(* Logix 5000 project; controller FV vendor 1 type 14 code 217 rev 31.11; software revision 31.00; part 19 of 63 *)
(* tags used below, declared in another part *)
   CheckTimeMask : INT;
   Delphi_Does_Eng_Func : BOOL;
   FR_FRV1_AV01 : PlantItem;   // FRV1_AV01
   FR_FV26_AV01 : PlantItem;   // FV26_AV01
   FR_FV26_AV04 : PlantItem;   // FV26_AV04
   FR_FV28_VA01 : PlantItem;   // FV28_VA01
   FR_FV29_VA01 : PlantItem;   // FV29_VA01
   FR_FV30_VA01 : PlantItem;   // FV30_VA01
   FR_FV31_VA01 : PlantItem;   // FV31_VA01
   FR_FVR1_P01 : PlantItem;   // FVR1_P01
   FR_FVS_P01 : PlantItem;   // FVS_P01
   FR_GBM_P01 : PlantItem;   // GBM_P01
   FR_N255 : INT[265];   // CHECKWORDS
   FR_YM_P01 : PlantItem;   // YM_P01
   FR_YM_P02 : PlantItem;   // YM_P02
   FR_YM_P03 : PlantItem;   // YM_P03
   TempChecktime : DINT;
(* FR_Common, continued *)

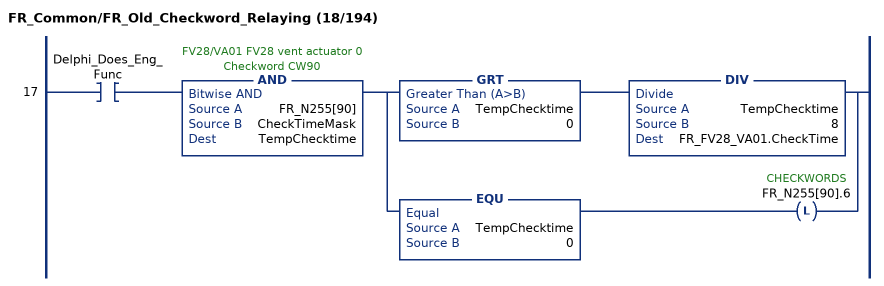
   [picture p322: FR_Common/FR_Old_Checkword_Relaying rungs 17-17]
   17: XIC(Delphi_Does_Eng_Func)AND(FR_N255[90],CheckTimeMask,TempChecktime)[GRT(TempChecktime,0) DIV(TempChecktime,8,FR_FV28_VA01.CheckTime) ,EQU(TempChecktime,0) OTL(FR_N255[90].6) ];
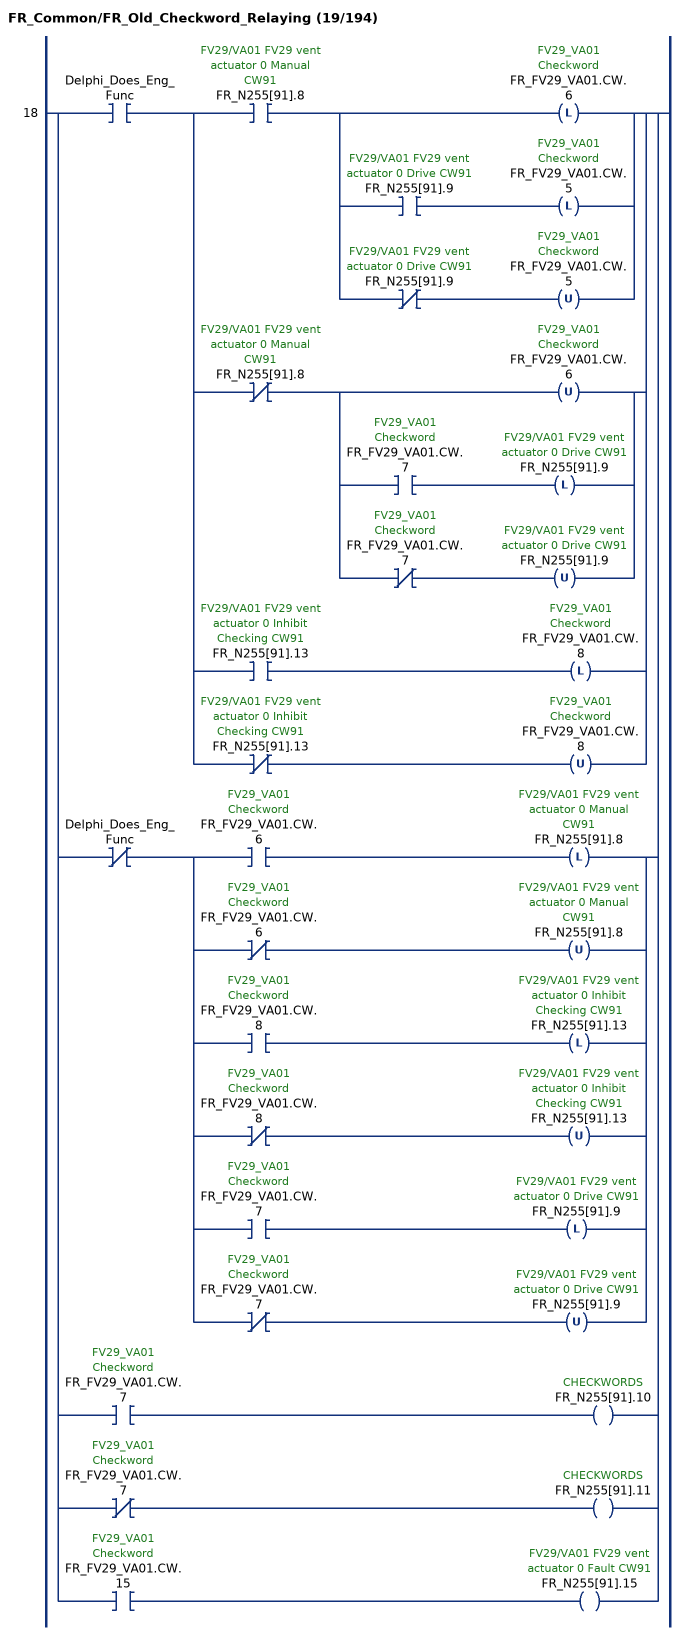
   18: [XIC(Delphi_Does_Eng_Func) [[XIC(FR_N255[91].8) [OTL(FR_FV29_VA01.CW.6) ,XIC(FR_N255[91].9) OTL(FR_FV29_VA01.CW.5) ,XIO(FR_N255[91].9) OTU(FR_FV29_VA01.CW.5) ] ,XIO(FR_N255[91].8) [OTU(FR_FV29_VA01.CW.6) ,[XIC(FR_FV29_VA01.CW.7) OTL(FR_N255[91].9) ,XIO(FR_FV29_VA01.CW.7) OTU(FR_N255[91].9) ] ] ] ,[XIC(FR_N255[91].13) OTL(FR_FV29_VA01.CW.8) ,XIO(FR_N255[91].13) OTU(FR_FV29_VA01.CW.8) ] ] ,XIO(Delphi_Does_Eng_Func) [[XIC(FR_FV29_VA01.CW.6) OTL(FR_N255[91].8) ,XIO(FR_FV29_VA01.CW.6) OTU(FR_N255[91].8) ] ,[XIC(FR_FV29_VA01.CW.8) OTL(FR_N255[91].13) ,XIO(FR_FV29_VA01.CW.8) OTU(FR_N255[91].13) ] ,[XIC(FR_FV29_VA01.CW.7) OTL(FR_N255[91].9) ,XIO(FR_FV29_VA01.CW.7) OTU(FR_N255[91].9) ] ] ,XIC(FR_FV29_VA01.CW.7) OTE(FR_N255[91].10) ,XIO(FR_FV29_VA01.CW.7) OTE(FR_N255[91].11) ,XIC(FR_FV29_VA01.CW.15) OTE(FR_N255[91].15) ];
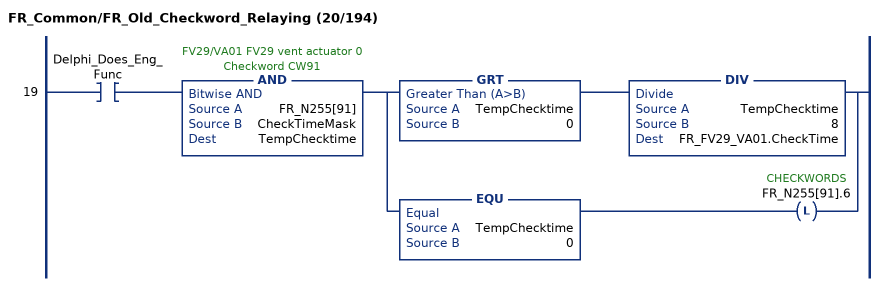
   19: XIC(Delphi_Does_Eng_Func)AND(FR_N255[91],CheckTimeMask,TempChecktime)[GRT(TempChecktime,0) DIV(TempChecktime,8,FR_FV29_VA01.CheckTime) ,EQU(TempChecktime,0) OTL(FR_N255[91].6) ];
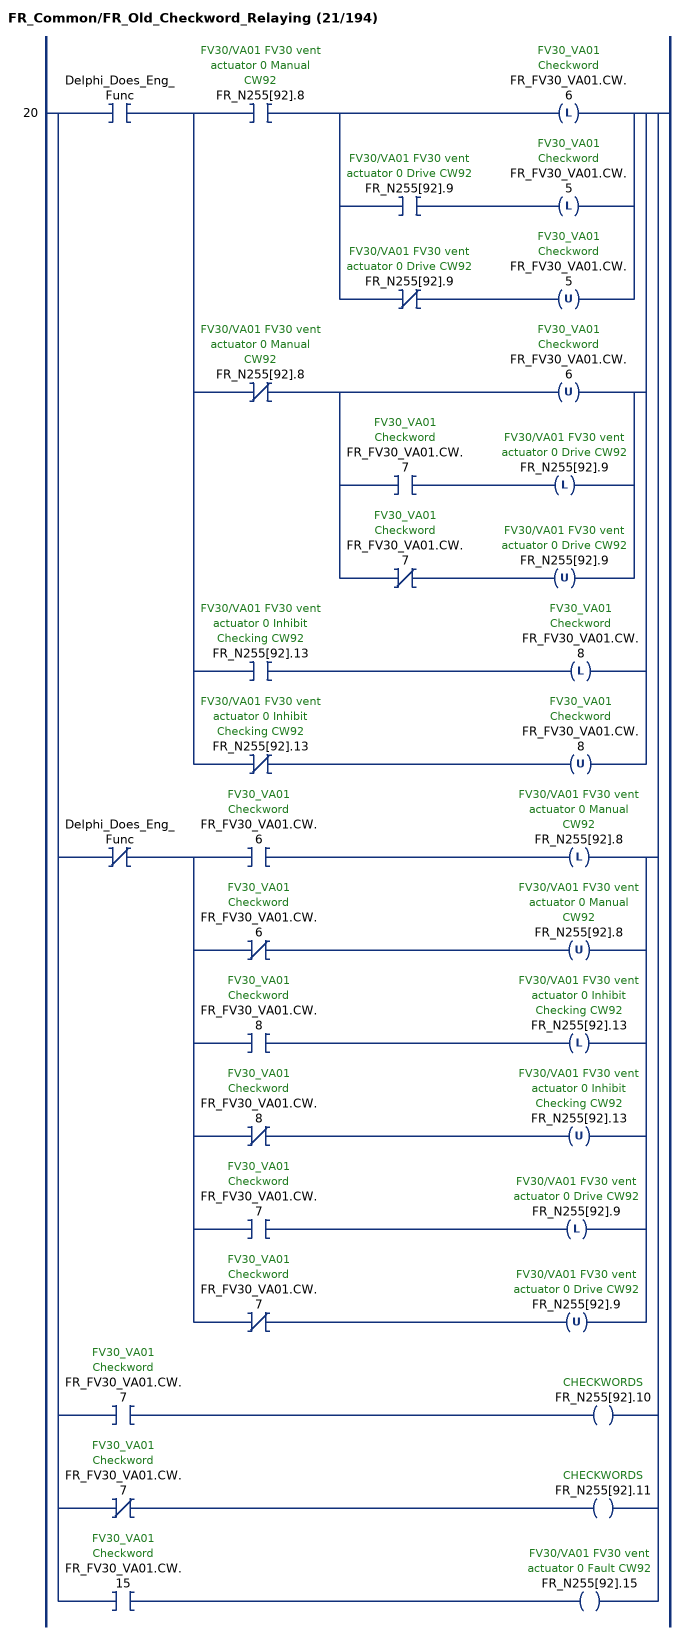
   20: [XIC(Delphi_Does_Eng_Func) [[XIC(FR_N255[92].8) [OTL(FR_FV30_VA01.CW.6) ,XIC(FR_N255[92].9) OTL(FR_FV30_VA01.CW.5) ,XIO(FR_N255[92].9) OTU(FR_FV30_VA01.CW.5) ] ,XIO(FR_N255[92].8) [OTU(FR_FV30_VA01.CW.6) ,[XIC(FR_FV30_VA01.CW.7) OTL(FR_N255[92].9) ,XIO(FR_FV30_VA01.CW.7) OTU(FR_N255[92].9) ] ] ] ,[XIC(FR_N255[92].13) OTL(FR_FV30_VA01.CW.8) ,XIO(FR_N255[92].13) OTU(FR_FV30_VA01.CW.8) ] ] ,XIO(Delphi_Does_Eng_Func) [[XIC(FR_FV30_VA01.CW.6) OTL(FR_N255[92].8) ,XIO(FR_FV30_VA01.CW.6) OTU(FR_N255[92].8) ] ,[XIC(FR_FV30_VA01.CW.8) OTL(FR_N255[92].13) ,XIO(FR_FV30_VA01.CW.8) OTU(FR_N255[92].13) ] ,[XIC(FR_FV30_VA01.CW.7) OTL(FR_N255[92].9) ,XIO(FR_FV30_VA01.CW.7) OTU(FR_N255[92].9) ] ] ,XIC(FR_FV30_VA01.CW.7) OTE(FR_N255[92].10) ,XIO(FR_FV30_VA01.CW.7) OTE(FR_N255[92].11) ,XIC(FR_FV30_VA01.CW.15) OTE(FR_N255[92].15) ];
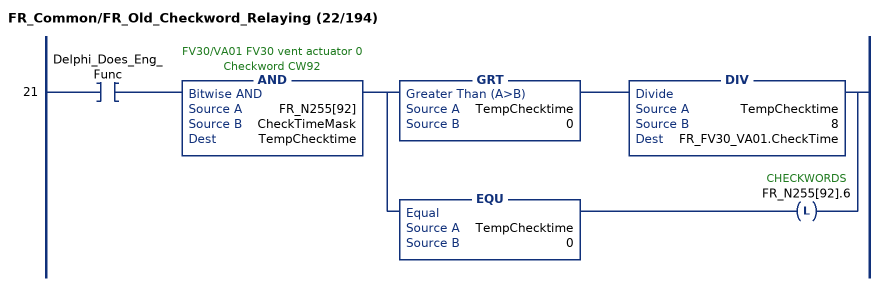
   21: XIC(Delphi_Does_Eng_Func)AND(FR_N255[92],CheckTimeMask,TempChecktime)[GRT(TempChecktime,0) DIV(TempChecktime,8,FR_FV30_VA01.CheckTime) ,EQU(TempChecktime,0) OTL(FR_N255[92].6) ];
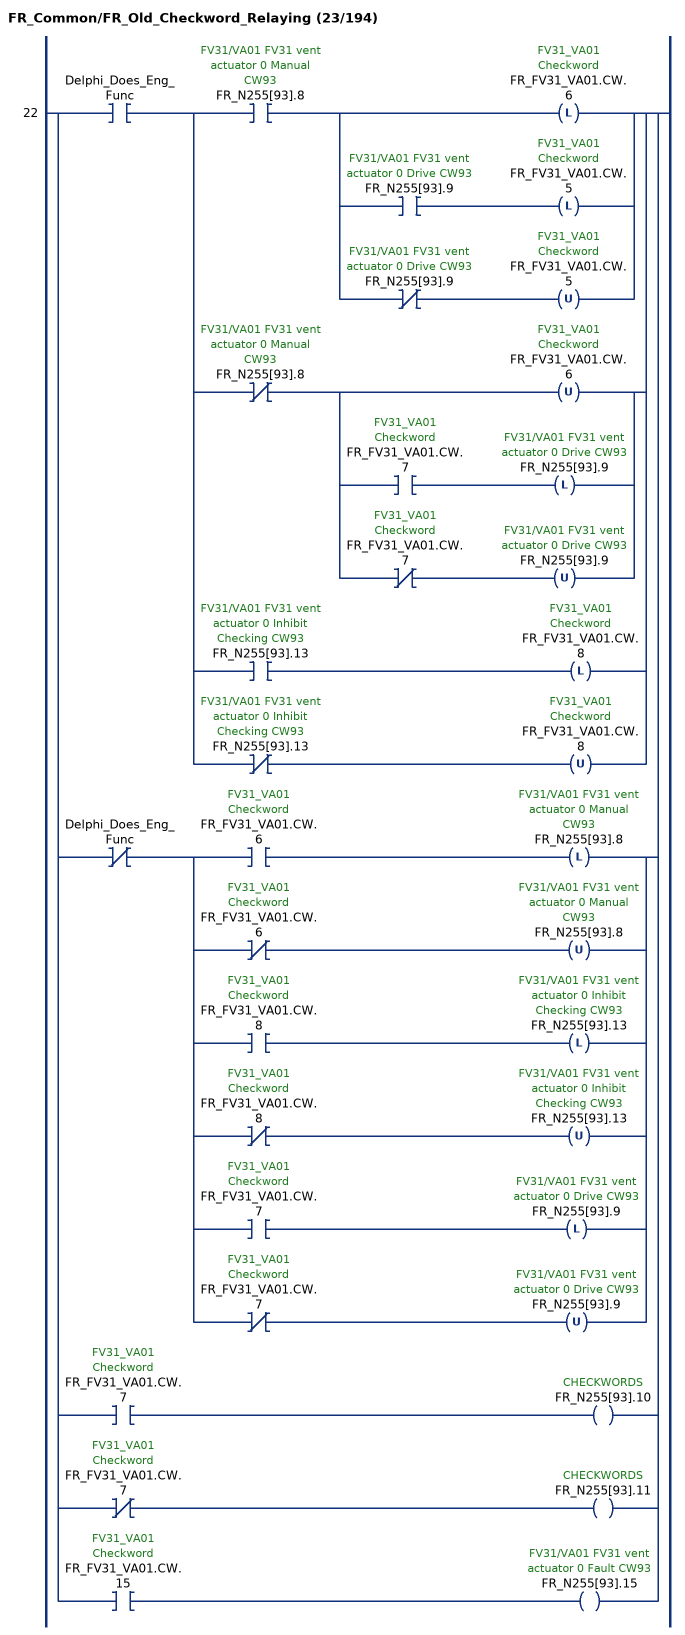
   22: [XIC(Delphi_Does_Eng_Func) [[XIC(FR_N255[93].8) [OTL(FR_FV31_VA01.CW.6) ,XIC(FR_N255[93].9) OTL(FR_FV31_VA01.CW.5) ,XIO(FR_N255[93].9) OTU(FR_FV31_VA01.CW.5) ] ,XIO(FR_N255[93].8) [OTU(FR_FV31_VA01.CW.6) ,[XIC(FR_FV31_VA01.CW.7) OTL(FR_N255[93].9) ,XIO(FR_FV31_VA01.CW.7) OTU(FR_N255[93].9) ] ] ] ,[XIC(FR_N255[93].13) OTL(FR_FV31_VA01.CW.8) ,XIO(FR_N255[93].13) OTU(FR_FV31_VA01.CW.8) ] ] ,XIO(Delphi_Does_Eng_Func) [[XIC(FR_FV31_VA01.CW.6) OTL(FR_N255[93].8) ,XIO(FR_FV31_VA01.CW.6) OTU(FR_N255[93].8) ] ,[XIC(FR_FV31_VA01.CW.8) OTL(FR_N255[93].13) ,XIO(FR_FV31_VA01.CW.8) OTU(FR_N255[93].13) ] ,[XIC(FR_FV31_VA01.CW.7) OTL(FR_N255[93].9) ,XIO(FR_FV31_VA01.CW.7) OTU(FR_N255[93].9) ] ] ,XIC(FR_FV31_VA01.CW.7) OTE(FR_N255[93].10) ,XIO(FR_FV31_VA01.CW.7) OTE(FR_N255[93].11) ,XIC(FR_FV31_VA01.CW.15) OTE(FR_N255[93].15) ];
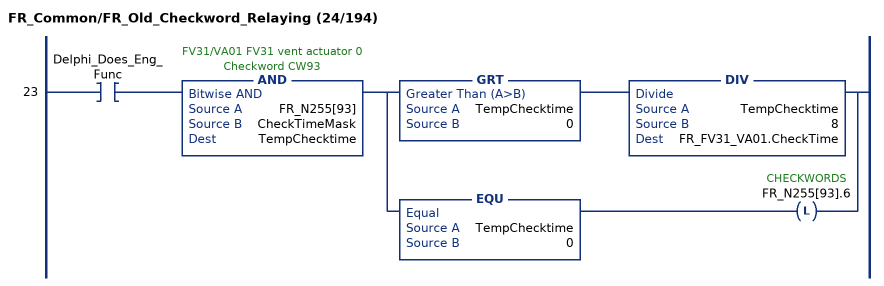
   23: XIC(Delphi_Does_Eng_Func)AND(FR_N255[93],CheckTimeMask,TempChecktime)[GRT(TempChecktime,0) DIV(TempChecktime,8,FR_FV31_VA01.CheckTime) ,EQU(TempChecktime,0) OTL(FR_N255[93].6) ];
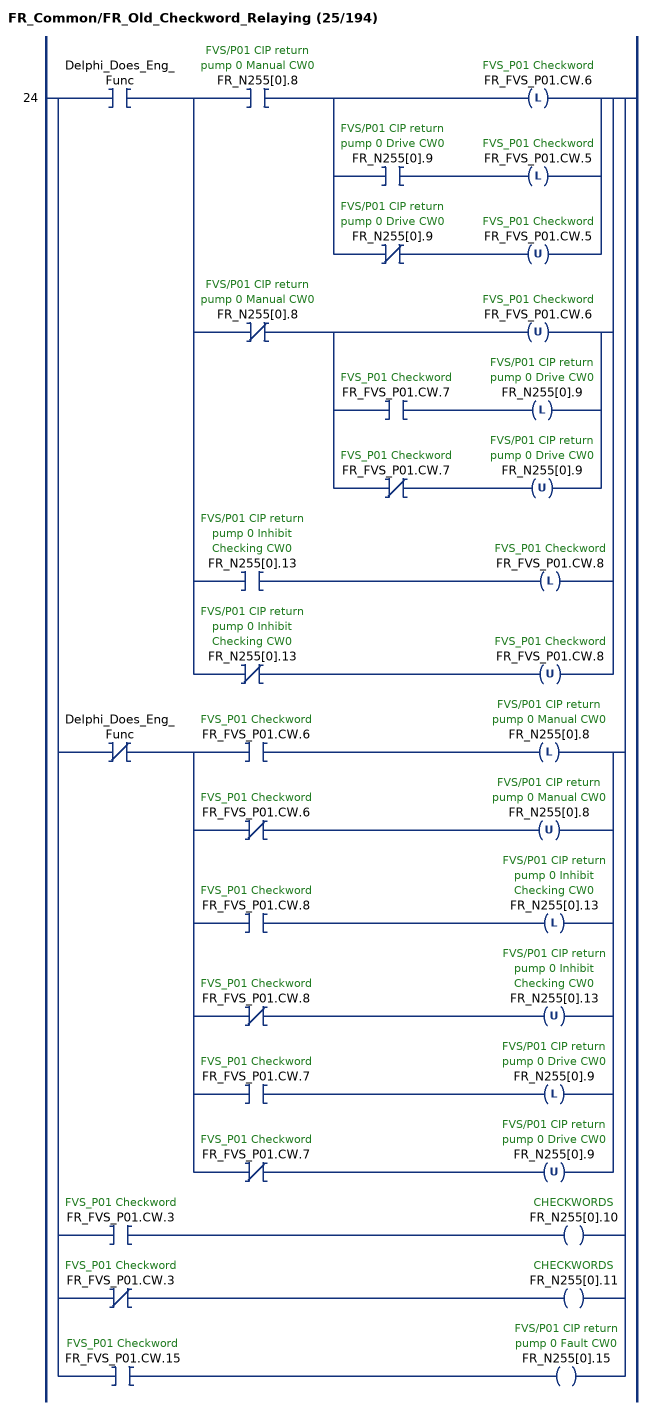
   24: [XIC(Delphi_Does_Eng_Func) [[XIC(FR_N255[0].8) [OTL(FR_FVS_P01.CW.6) ,XIC(FR_N255[0].9) OTL(FR_FVS_P01.CW.5) ,XIO(FR_N255[0].9) OTU(FR_FVS_P01.CW.5) ] ,XIO(FR_N255[0].8) [OTU(FR_FVS_P01.CW.6) ,[XIC(FR_FVS_P01.CW.7) OTL(FR_N255[0].9) ,XIO(FR_FVS_P01.CW.7) OTU(FR_N255[0].9) ] ] ] ,[XIC(FR_N255[0].13) OTL(FR_FVS_P01.CW.8) ,XIO(FR_N255[0].13) OTU(FR_FVS_P01.CW.8) ] ] ,XIO(Delphi_Does_Eng_Func) [[XIC(FR_FVS_P01.CW.6) OTL(FR_N255[0].8) ,XIO(FR_FVS_P01.CW.6) OTU(FR_N255[0].8) ] ,[XIC(FR_FVS_P01.CW.8) OTL(FR_N255[0].13) ,XIO(FR_FVS_P01.CW.8) OTU(FR_N255[0].13) ] ,[XIC(FR_FVS_P01.CW.7) OTL(FR_N255[0].9) ,XIO(FR_FVS_P01.CW.7) OTU(FR_N255[0].9) ] ] ,XIC(FR_FVS_P01.CW.3) OTE(FR_N255[0].10) ,XIO(FR_FVS_P01.CW.3) OTE(FR_N255[0].11) ,XIC(FR_FVS_P01.CW.15) OTE(FR_N255[0].15) ];
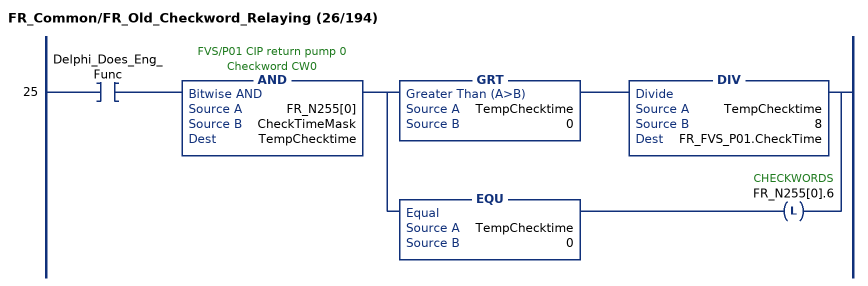
   25: XIC(Delphi_Does_Eng_Func)AND(FR_N255[0],CheckTimeMask,TempChecktime)[GRT(TempChecktime,0) DIV(TempChecktime,8,FR_FVS_P01.CheckTime) ,EQU(TempChecktime,0) OTL(FR_N255[0].6) ];
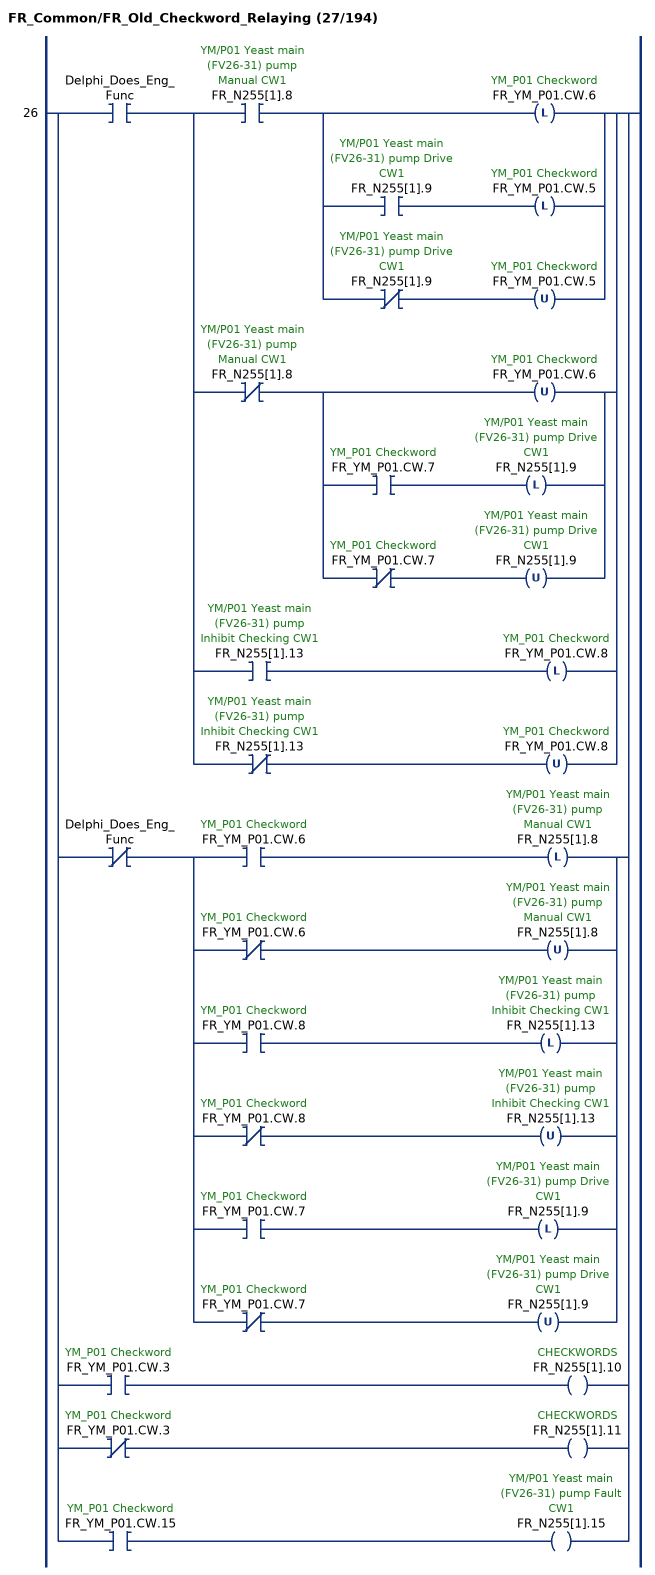
   26: [XIC(Delphi_Does_Eng_Func) [[XIC(FR_N255[1].8) [OTL(FR_YM_P01.CW.6) ,XIC(FR_N255[1].9) OTL(FR_YM_P01.CW.5) ,XIO(FR_N255[1].9) OTU(FR_YM_P01.CW.5) ] ,XIO(FR_N255[1].8) [OTU(FR_YM_P01.CW.6) ,[XIC(FR_YM_P01.CW.7) OTL(FR_N255[1].9) ,XIO(FR_YM_P01.CW.7) OTU(FR_N255[1].9) ] ] ] ,[XIC(FR_N255[1].13) OTL(FR_YM_P01.CW.8) ,XIO(FR_N255[1].13) OTU(FR_YM_P01.CW.8) ] ] ,XIO(Delphi_Does_Eng_Func) [[XIC(FR_YM_P01.CW.6) OTL(FR_N255[1].8) ,XIO(FR_YM_P01.CW.6) OTU(FR_N255[1].8) ] ,[XIC(FR_YM_P01.CW.8) OTL(FR_N255[1].13) ,XIO(FR_YM_P01.CW.8) OTU(FR_N255[1].13) ] ,[XIC(FR_YM_P01.CW.7) OTL(FR_N255[1].9) ,XIO(FR_YM_P01.CW.7) OTU(FR_N255[1].9) ] ] ,XIC(FR_YM_P01.CW.3) OTE(FR_N255[1].10) ,XIO(FR_YM_P01.CW.3) OTE(FR_N255[1].11) ,XIC(FR_YM_P01.CW.15) OTE(FR_N255[1].15) ];
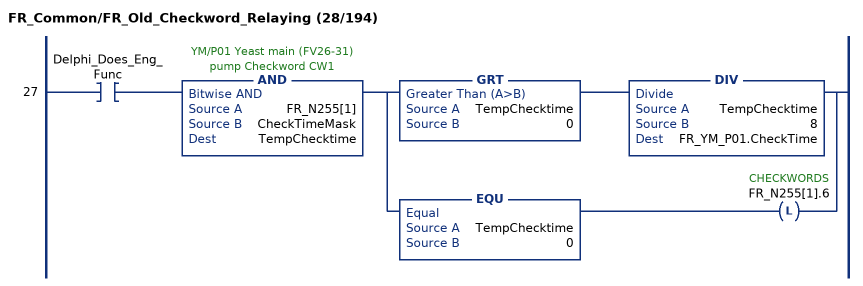
   27: XIC(Delphi_Does_Eng_Func)AND(FR_N255[1],CheckTimeMask,TempChecktime)[GRT(TempChecktime,0) DIV(TempChecktime,8,FR_YM_P01.CheckTime) ,EQU(TempChecktime,0) OTL(FR_N255[1].6) ];
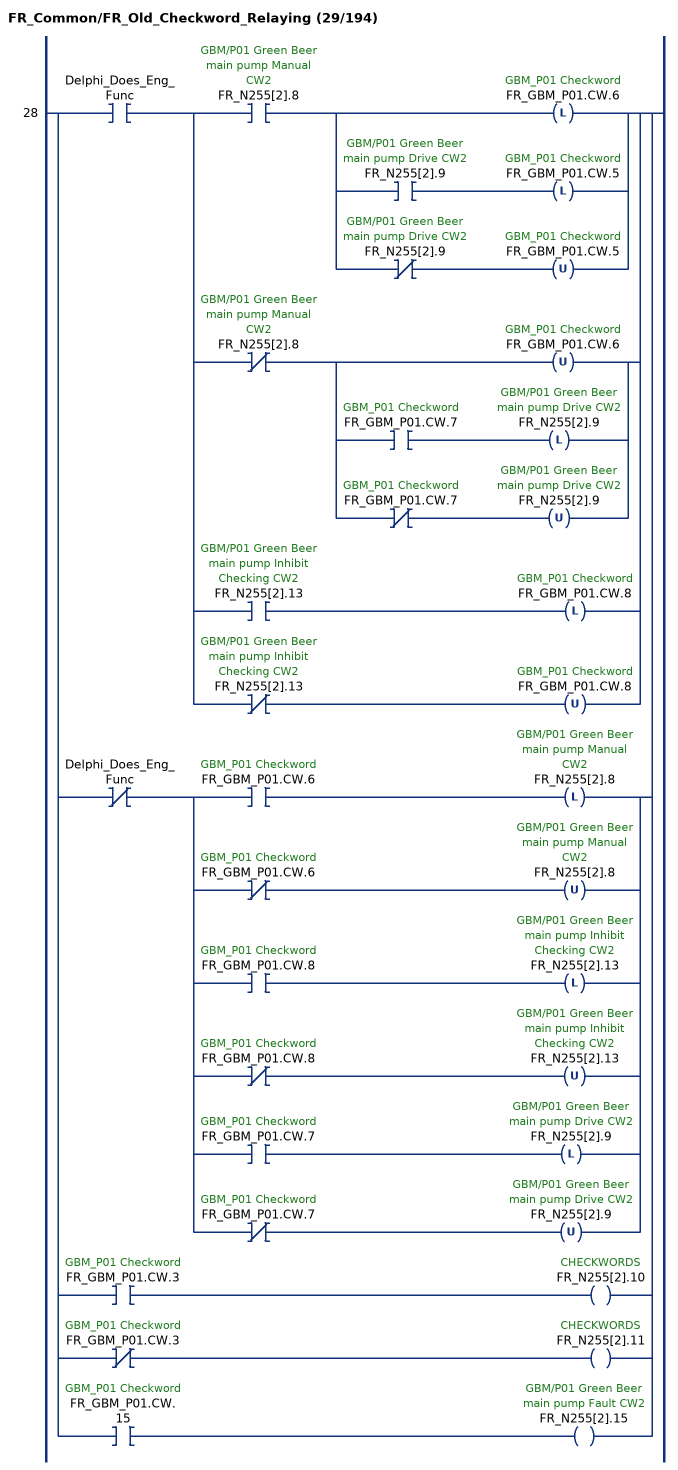
   28: [XIC(Delphi_Does_Eng_Func) [[XIC(FR_N255[2].8) [OTL(FR_GBM_P01.CW.6) ,XIC(FR_N255[2].9) OTL(FR_GBM_P01.CW.5) ,XIO(FR_N255[2].9) OTU(FR_GBM_P01.CW.5) ] ,XIO(FR_N255[2].8) [OTU(FR_GBM_P01.CW.6) ,[XIC(FR_GBM_P01.CW.7) OTL(FR_N255[2].9) ,XIO(FR_GBM_P01.CW.7) OTU(FR_N255[2].9) ] ] ] ,[XIC(FR_N255[2].13) OTL(FR_GBM_P01.CW.8) ,XIO(FR_N255[2].13) OTU(FR_GBM_P01.CW.8) ] ] ,XIO(Delphi_Does_Eng_Func) [[XIC(FR_GBM_P01.CW.6) OTL(FR_N255[2].8) ,XIO(FR_GBM_P01.CW.6) OTU(FR_N255[2].8) ] ,[XIC(FR_GBM_P01.CW.8) OTL(FR_N255[2].13) ,XIO(FR_GBM_P01.CW.8) OTU(FR_N255[2].13) ] ,[XIC(FR_GBM_P01.CW.7) OTL(FR_N255[2].9) ,XIO(FR_GBM_P01.CW.7) OTU(FR_N255[2].9) ] ] ,XIC(FR_GBM_P01.CW.3) OTE(FR_N255[2].10) ,XIO(FR_GBM_P01.CW.3) OTE(FR_N255[2].11) ,XIC(FR_GBM_P01.CW.15) OTE(FR_N255[2].15) ];
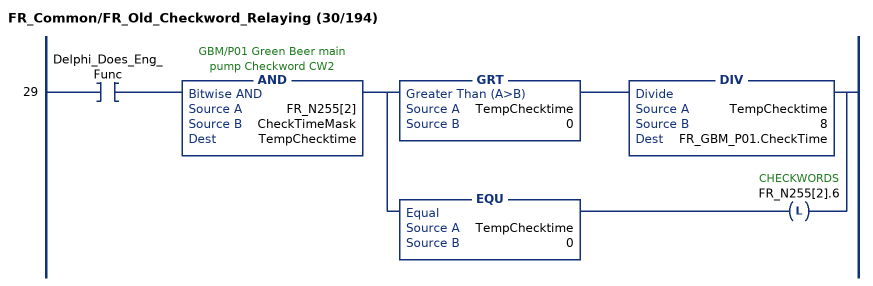
   29: XIC(Delphi_Does_Eng_Func)AND(FR_N255[2],CheckTimeMask,TempChecktime)[GRT(TempChecktime,0) DIV(TempChecktime,8,FR_GBM_P01.CheckTime) ,EQU(TempChecktime,0) OTL(FR_N255[2].6) ];
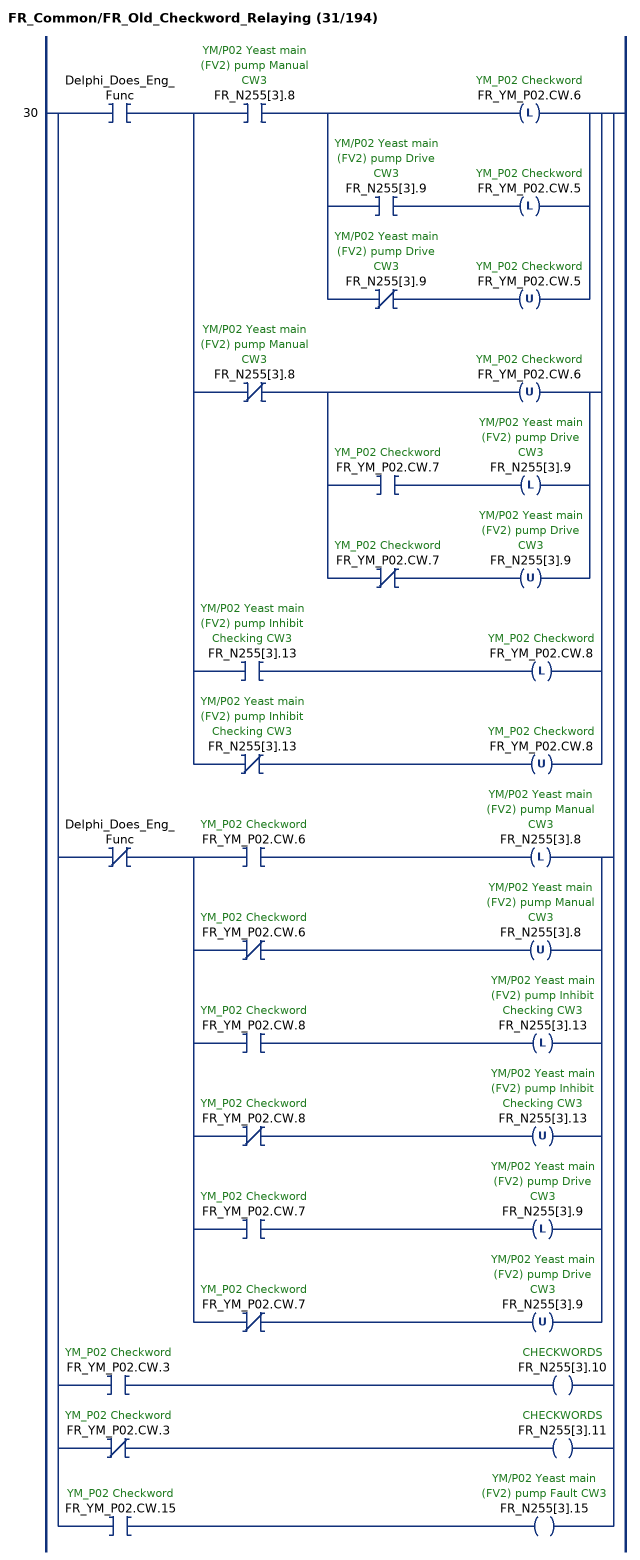
   30: [XIC(Delphi_Does_Eng_Func) [[XIC(FR_N255[3].8) [OTL(FR_YM_P02.CW.6) ,XIC(FR_N255[3].9) OTL(FR_YM_P02.CW.5) ,XIO(FR_N255[3].9) OTU(FR_YM_P02.CW.5) ] ,XIO(FR_N255[3].8) [OTU(FR_YM_P02.CW.6) ,[XIC(FR_YM_P02.CW.7) OTL(FR_N255[3].9) ,XIO(FR_YM_P02.CW.7) OTU(FR_N255[3].9) ] ] ] ,[XIC(FR_N255[3].13) OTL(FR_YM_P02.CW.8) ,XIO(FR_N255[3].13) OTU(FR_YM_P02.CW.8) ] ] ,XIO(Delphi_Does_Eng_Func) [[XIC(FR_YM_P02.CW.6) OTL(FR_N255[3].8) ,XIO(FR_YM_P02.CW.6) OTU(FR_N255[3].8) ] ,[XIC(FR_YM_P02.CW.8) OTL(FR_N255[3].13) ,XIO(FR_YM_P02.CW.8) OTU(FR_N255[3].13) ] ,[XIC(FR_YM_P02.CW.7) OTL(FR_N255[3].9) ,XIO(FR_YM_P02.CW.7) OTU(FR_N255[3].9) ] ] ,XIC(FR_YM_P02.CW.3) OTE(FR_N255[3].10) ,XIO(FR_YM_P02.CW.3) OTE(FR_N255[3].11) ,XIC(FR_YM_P02.CW.15) OTE(FR_N255[3].15) ];
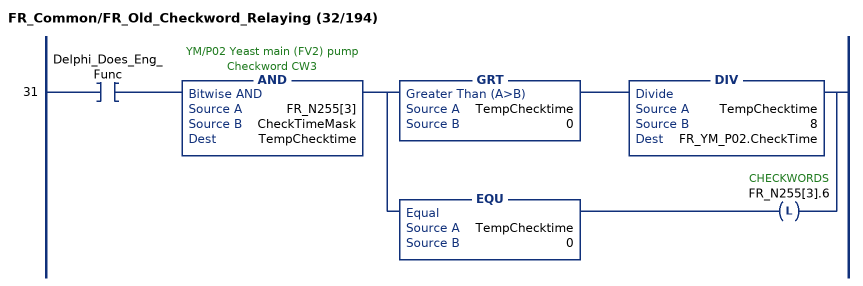
   31: XIC(Delphi_Does_Eng_Func)AND(FR_N255[3],CheckTimeMask,TempChecktime)[GRT(TempChecktime,0) DIV(TempChecktime,8,FR_YM_P02.CheckTime) ,EQU(TempChecktime,0) OTL(FR_N255[3].6) ];
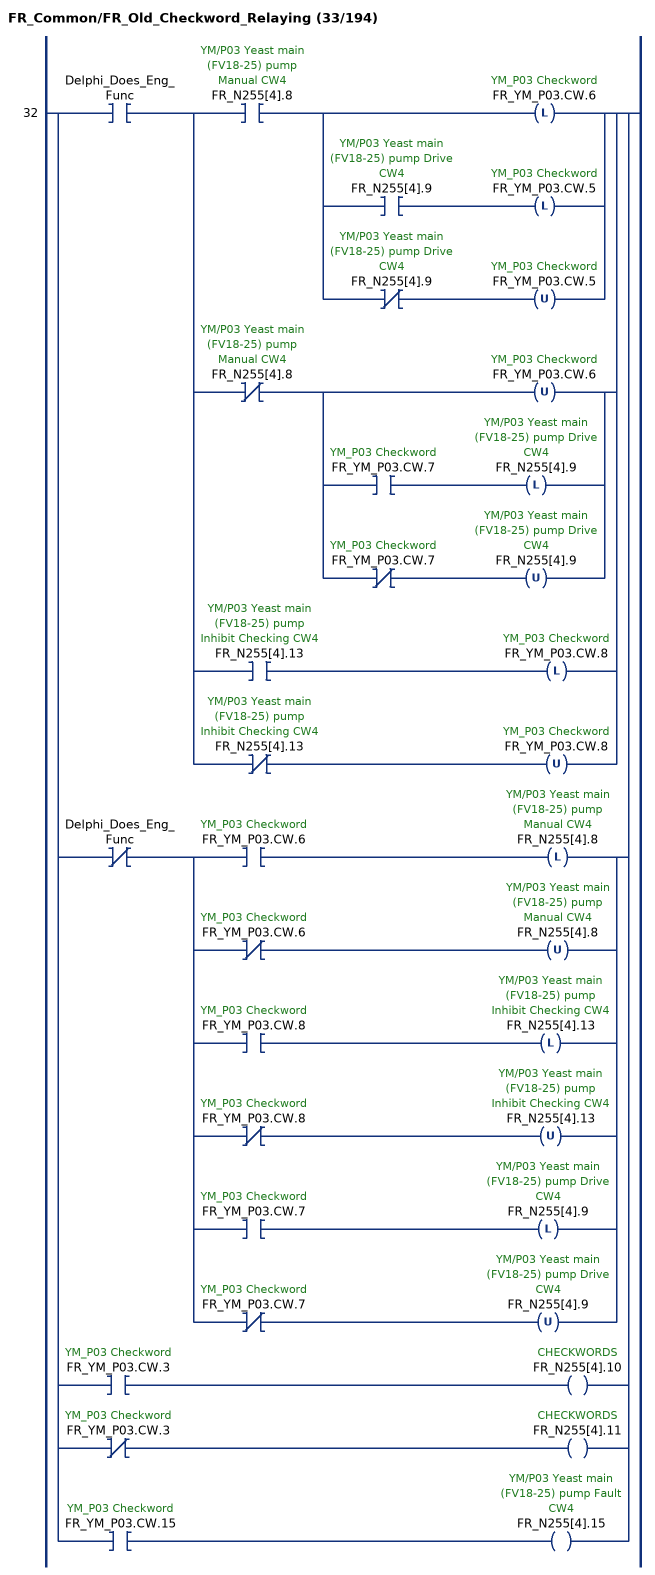
   32: [XIC(Delphi_Does_Eng_Func) [[XIC(FR_N255[4].8) [OTL(FR_YM_P03.CW.6) ,XIC(FR_N255[4].9) OTL(FR_YM_P03.CW.5) ,XIO(FR_N255[4].9) OTU(FR_YM_P03.CW.5) ] ,XIO(FR_N255[4].8) [OTU(FR_YM_P03.CW.6) ,[XIC(FR_YM_P03.CW.7) OTL(FR_N255[4].9) ,XIO(FR_YM_P03.CW.7) OTU(FR_N255[4].9) ] ] ] ,[XIC(FR_N255[4].13) OTL(FR_YM_P03.CW.8) ,XIO(FR_N255[4].13) OTU(FR_YM_P03.CW.8) ] ] ,XIO(Delphi_Does_Eng_Func) [[XIC(FR_YM_P03.CW.6) OTL(FR_N255[4].8) ,XIO(FR_YM_P03.CW.6) OTU(FR_N255[4].8) ] ,[XIC(FR_YM_P03.CW.8) OTL(FR_N255[4].13) ,XIO(FR_YM_P03.CW.8) OTU(FR_N255[4].13) ] ,[XIC(FR_YM_P03.CW.7) OTL(FR_N255[4].9) ,XIO(FR_YM_P03.CW.7) OTU(FR_N255[4].9) ] ] ,XIC(FR_YM_P03.CW.3) OTE(FR_N255[4].10) ,XIO(FR_YM_P03.CW.3) OTE(FR_N255[4].11) ,XIC(FR_YM_P03.CW.15) OTE(FR_N255[4].15) ];
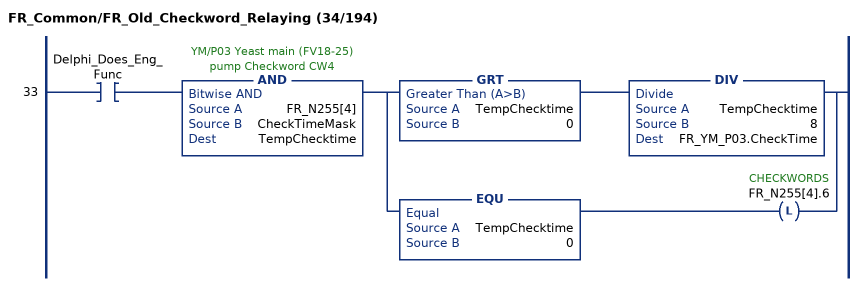
   33: XIC(Delphi_Does_Eng_Func)AND(FR_N255[4],CheckTimeMask,TempChecktime)[GRT(TempChecktime,0) DIV(TempChecktime,8,FR_YM_P03.CheckTime) ,EQU(TempChecktime,0) OTL(FR_N255[4].6) ];
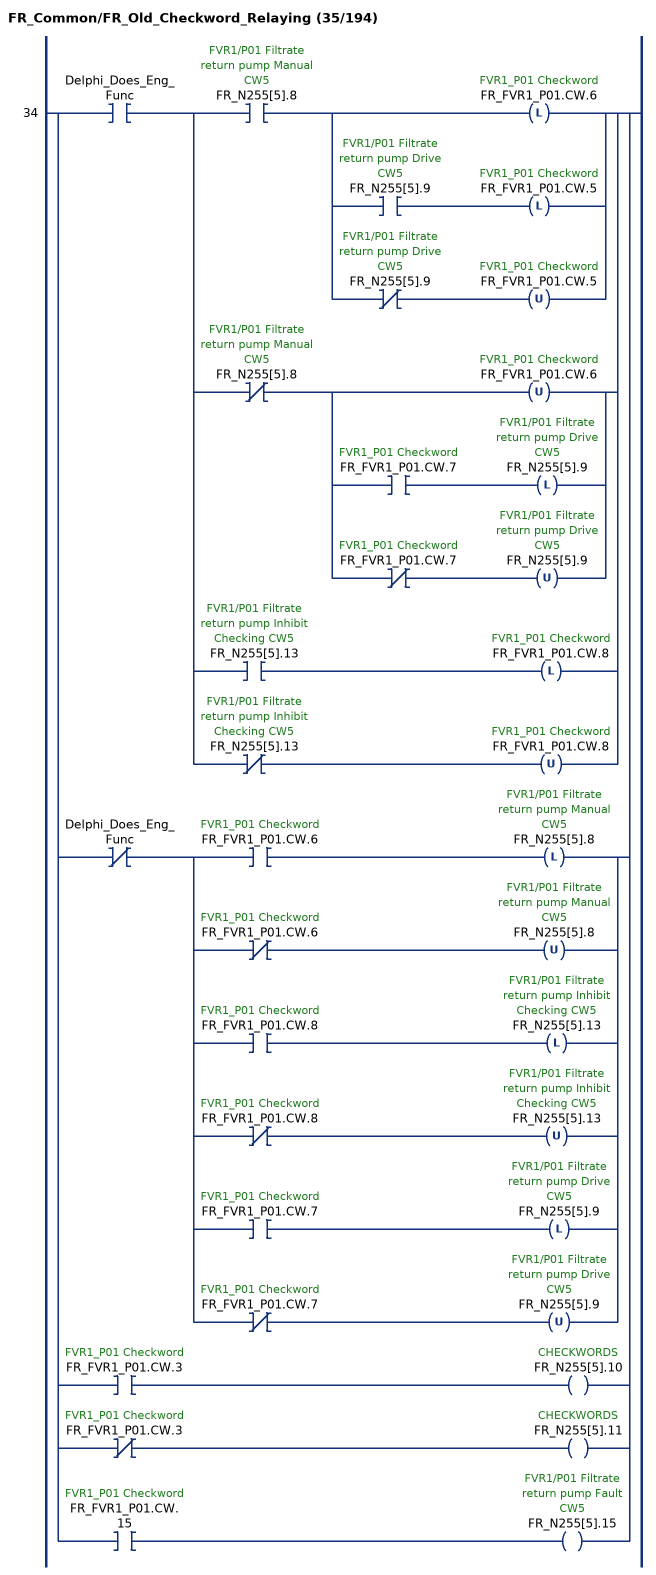
   34: [XIC(Delphi_Does_Eng_Func) [[XIC(FR_N255[5].8) [OTL(FR_FVR1_P01.CW.6) ,XIC(FR_N255[5].9) OTL(FR_FVR1_P01.CW.5) ,XIO(FR_N255[5].9) OTU(FR_FVR1_P01.CW.5) ] ,XIO(FR_N255[5].8) [OTU(FR_FVR1_P01.CW.6) ,[XIC(FR_FVR1_P01.CW.7) OTL(FR_N255[5].9) ,XIO(FR_FVR1_P01.CW.7) OTU(FR_N255[5].9) ] ] ] ,[XIC(FR_N255[5].13) OTL(FR_FVR1_P01.CW.8) ,XIO(FR_N255[5].13) OTU(FR_FVR1_P01.CW.8) ] ] ,XIO(Delphi_Does_Eng_Func) [[XIC(FR_FVR1_P01.CW.6) OTL(FR_N255[5].8) ,XIO(FR_FVR1_P01.CW.6) OTU(FR_N255[5].8) ] ,[XIC(FR_FVR1_P01.CW.8) OTL(FR_N255[5].13) ,XIO(FR_FVR1_P01.CW.8) OTU(FR_N255[5].13) ] ,[XIC(FR_FVR1_P01.CW.7) OTL(FR_N255[5].9) ,XIO(FR_FVR1_P01.CW.7) OTU(FR_N255[5].9) ] ] ,XIC(FR_FVR1_P01.CW.3) OTE(FR_N255[5].10) ,XIO(FR_FVR1_P01.CW.3) OTE(FR_N255[5].11) ,XIC(FR_FVR1_P01.CW.15) OTE(FR_N255[5].15) ];
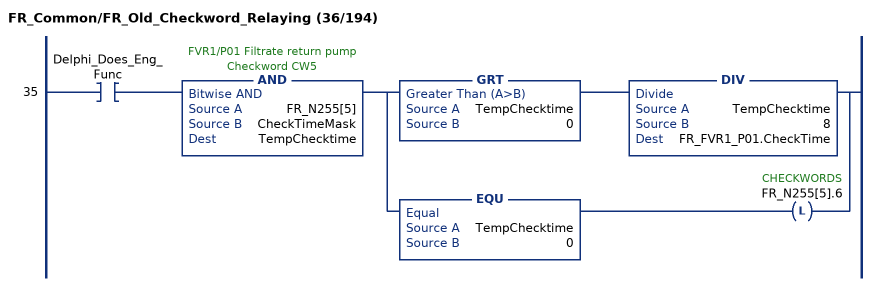
   35: XIC(Delphi_Does_Eng_Func)AND(FR_N255[5],CheckTimeMask,TempChecktime)[GRT(TempChecktime,0) DIV(TempChecktime,8,FR_FVR1_P01.CheckTime) ,EQU(TempChecktime,0) OTL(FR_N255[5].6) ];
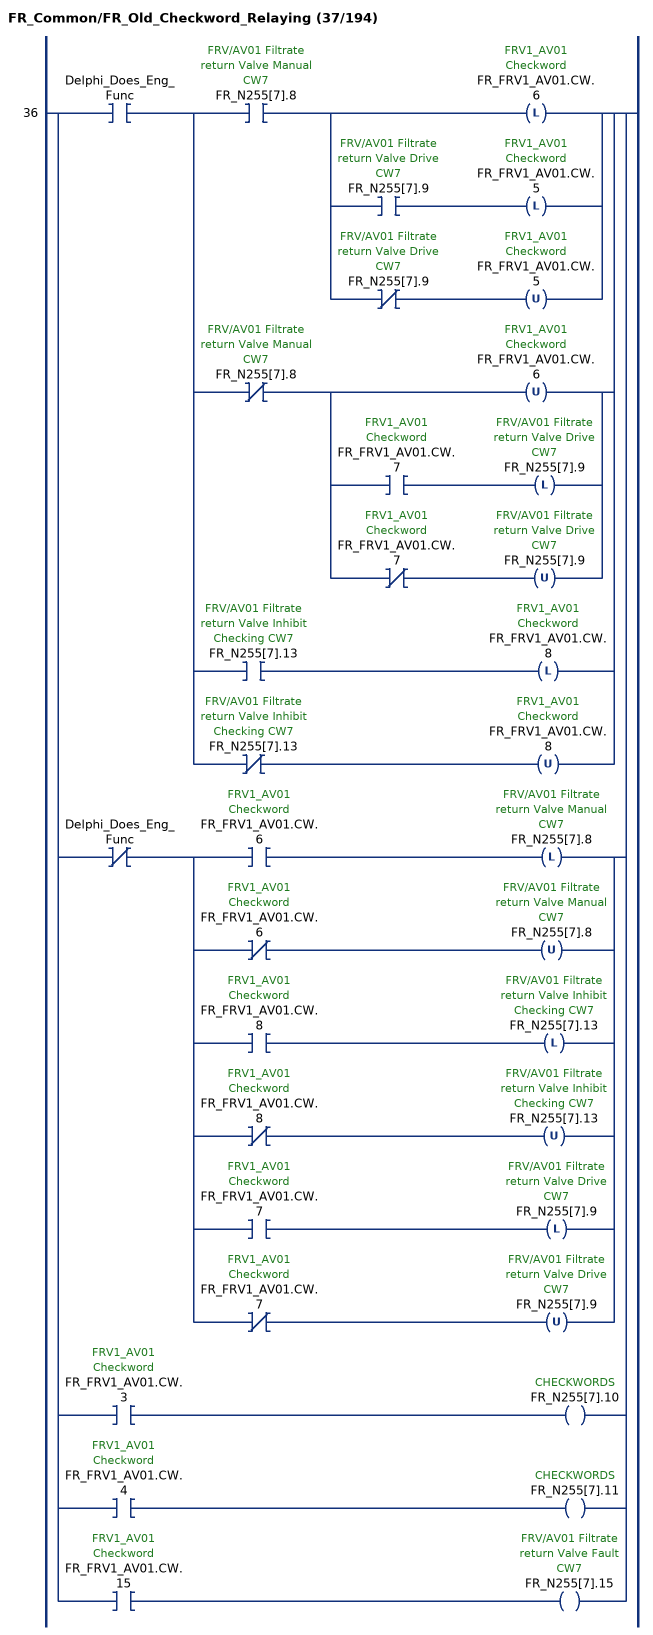
   36: [XIC(Delphi_Does_Eng_Func) [[XIC(FR_N255[7].8) [OTL(FR_FRV1_AV01.CW.6) ,XIC(FR_N255[7].9) OTL(FR_FRV1_AV01.CW.5) ,XIO(FR_N255[7].9) OTU(FR_FRV1_AV01.CW.5) ] ,XIO(FR_N255[7].8) [OTU(FR_FRV1_AV01.CW.6) ,[XIC(FR_FRV1_AV01.CW.7) OTL(FR_N255[7].9) ,XIO(FR_FRV1_AV01.CW.7) OTU(FR_N255[7].9) ] ] ] ,[XIC(FR_N255[7].13) OTL(FR_FRV1_AV01.CW.8) ,XIO(FR_N255[7].13) OTU(FR_FRV1_AV01.CW.8) ] ] ,XIO(Delphi_Does_Eng_Func) [[XIC(FR_FRV1_AV01.CW.6) OTL(FR_N255[7].8) ,XIO(FR_FRV1_AV01.CW.6) OTU(FR_N255[7].8) ] ,[XIC(FR_FRV1_AV01.CW.8) OTL(FR_N255[7].13) ,XIO(FR_FRV1_AV01.CW.8) OTU(FR_N255[7].13) ] ,[XIC(FR_FRV1_AV01.CW.7) OTL(FR_N255[7].9) ,XIO(FR_FRV1_AV01.CW.7) OTU(FR_N255[7].9) ] ] ,XIC(FR_FRV1_AV01.CW.3) OTE(FR_N255[7].10) ,XIC(FR_FRV1_AV01.CW.4) OTE(FR_N255[7].11) ,XIC(FR_FRV1_AV01.CW.15) OTE(FR_N255[7].15) ];
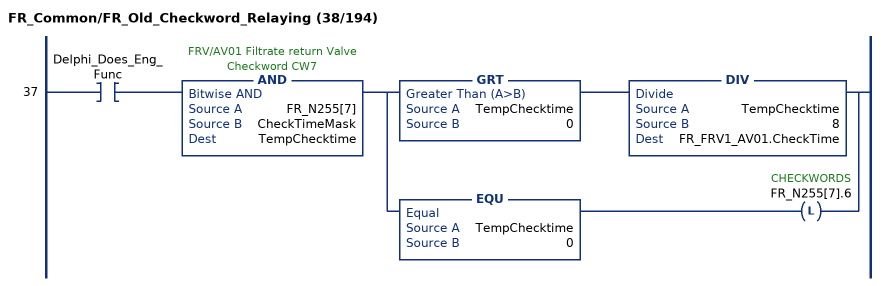
   37: XIC(Delphi_Does_Eng_Func)AND(FR_N255[7],CheckTimeMask,TempChecktime)[GRT(TempChecktime,0) DIV(TempChecktime,8,FR_FRV1_AV01.CheckTime) ,EQU(TempChecktime,0) OTL(FR_N255[7].6) ];
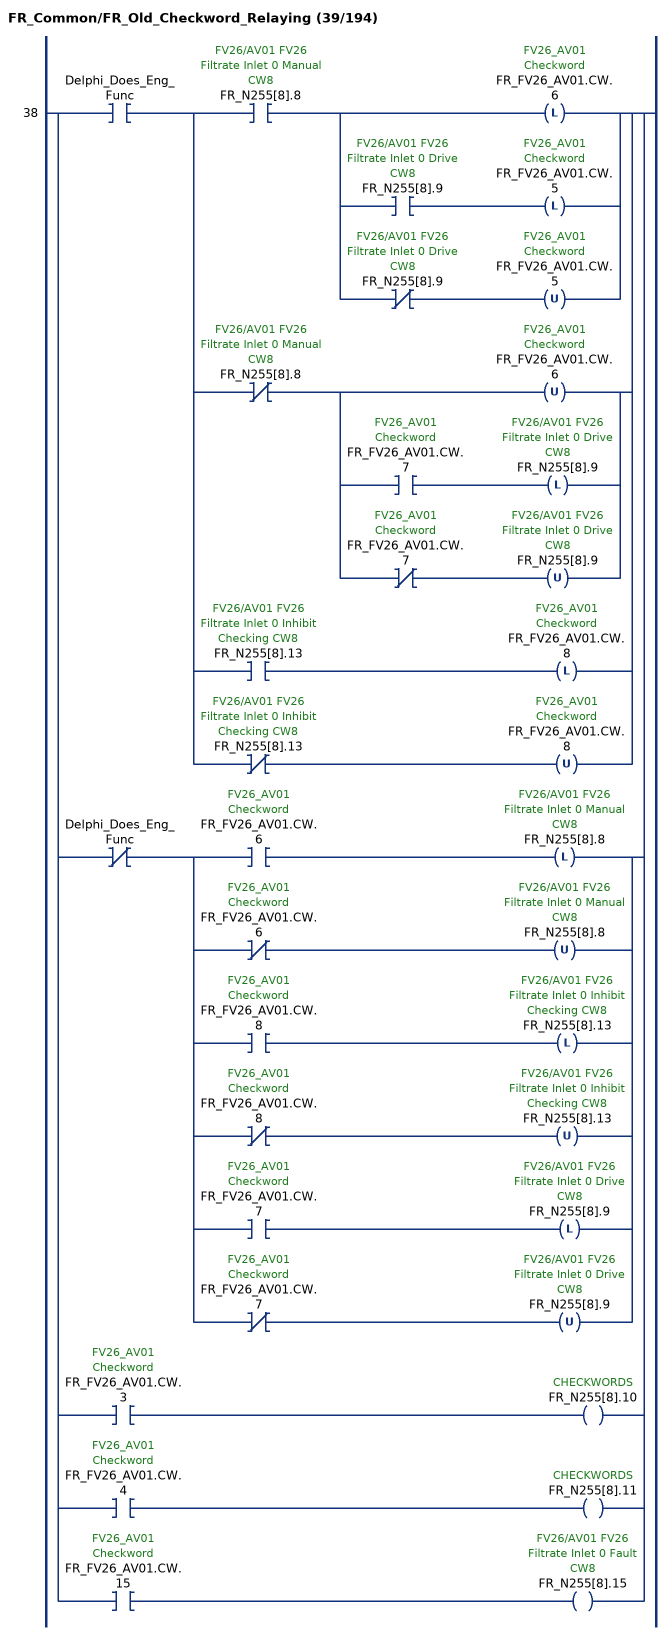
   38: [XIC(Delphi_Does_Eng_Func) [[XIC(FR_N255[8].8) [OTL(FR_FV26_AV01.CW.6) ,XIC(FR_N255[8].9) OTL(FR_FV26_AV01.CW.5) ,XIO(FR_N255[8].9) OTU(FR_FV26_AV01.CW.5) ] ,XIO(FR_N255[8].8) [OTU(FR_FV26_AV01.CW.6) ,[XIC(FR_FV26_AV01.CW.7) OTL(FR_N255[8].9) ,XIO(FR_FV26_AV01.CW.7) OTU(FR_N255[8].9) ] ] ] ,[XIC(FR_N255[8].13) OTL(FR_FV26_AV01.CW.8) ,XIO(FR_N255[8].13) OTU(FR_FV26_AV01.CW.8) ] ] ,XIO(Delphi_Does_Eng_Func) [[XIC(FR_FV26_AV01.CW.6) OTL(FR_N255[8].8) ,XIO(FR_FV26_AV01.CW.6) OTU(FR_N255[8].8) ] ,[XIC(FR_FV26_AV01.CW.8) OTL(FR_N255[8].13) ,XIO(FR_FV26_AV01.CW.8) OTU(FR_N255[8].13) ] ,[XIC(FR_FV26_AV01.CW.7) OTL(FR_N255[8].9) ,XIO(FR_FV26_AV01.CW.7) OTU(FR_N255[8].9) ] ] ,XIC(FR_FV26_AV01.CW.3) OTE(FR_N255[8].10) ,XIC(FR_FV26_AV01.CW.4) OTE(FR_N255[8].11) ,XIC(FR_FV26_AV01.CW.15) OTE(FR_N255[8].15) ];
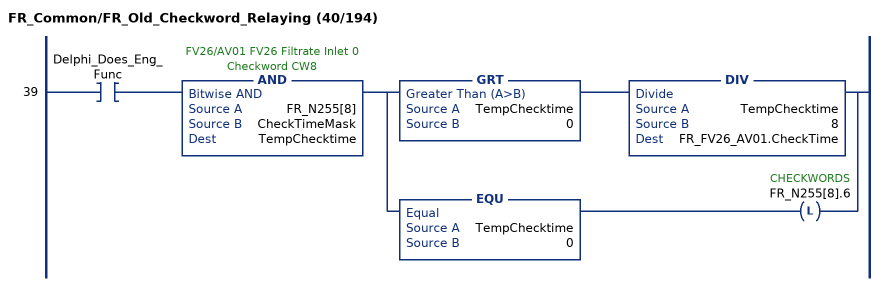
   39: XIC(Delphi_Does_Eng_Func)AND(FR_N255[8],CheckTimeMask,TempChecktime)[GRT(TempChecktime,0) DIV(TempChecktime,8,FR_FV26_AV01.CheckTime) ,EQU(TempChecktime,0) OTL(FR_N255[8].6) ];
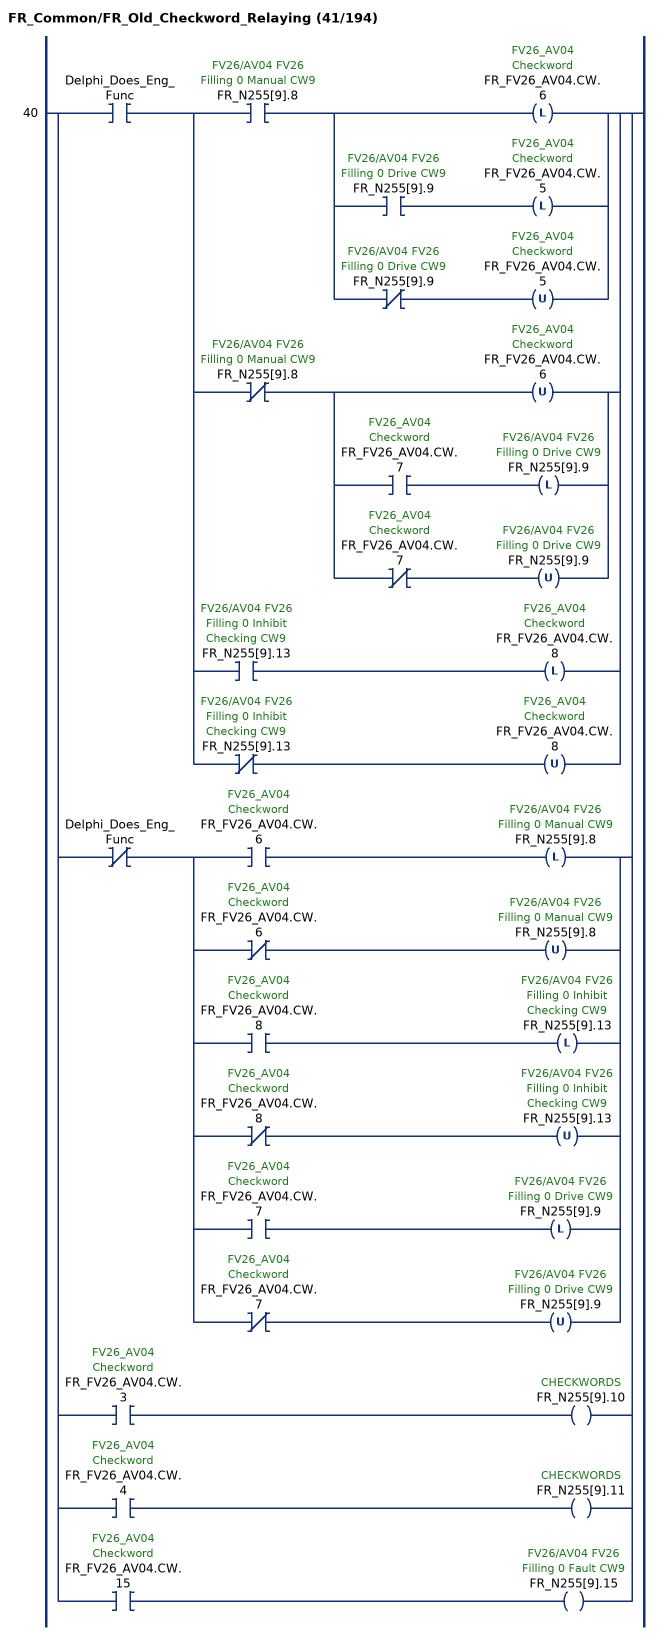
   40: [XIC(Delphi_Does_Eng_Func) [[XIC(FR_N255[9].8) [OTL(FR_FV26_AV04.CW.6) ,XIC(FR_N255[9].9) OTL(FR_FV26_AV04.CW.5) ,XIO(FR_N255[9].9) OTU(FR_FV26_AV04.CW.5) ] ,XIO(FR_N255[9].8) [OTU(FR_FV26_AV04.CW.6) ,[XIC(FR_FV26_AV04.CW.7) OTL(FR_N255[9].9) ,XIO(FR_FV26_AV04.CW.7) OTU(FR_N255[9].9) ] ] ] ,[XIC(FR_N255[9].13) OTL(FR_FV26_AV04.CW.8) ,XIO(FR_N255[9].13) OTU(FR_FV26_AV04.CW.8) ] ] ,XIO(Delphi_Does_Eng_Func) [[XIC(FR_FV26_AV04.CW.6) OTL(FR_N255[9].8) ,XIO(FR_FV26_AV04.CW.6) OTU(FR_N255[9].8) ] ,[XIC(FR_FV26_AV04.CW.8) OTL(FR_N255[9].13) ,XIO(FR_FV26_AV04.CW.8) OTU(FR_N255[9].13) ] ,[XIC(FR_FV26_AV04.CW.7) OTL(FR_N255[9].9) ,XIO(FR_FV26_AV04.CW.7) OTU(FR_N255[9].9) ] ] ,XIC(FR_FV26_AV04.CW.3) OTE(FR_N255[9].10) ,XIC(FR_FV26_AV04.CW.4) OTE(FR_N255[9].11) ,XIC(FR_FV26_AV04.CW.15) OTE(FR_N255[9].15) ];
